(* Logix 5000 project; controller Joltek_RA_5069PLC002 vendor 1 type 14 code 226 rev 34.15; software revision 34.04 *)

TASK MainTask (continuous, watchdog 500 ms) : MainProgram
TASK SafetyTask (periodic, rate 20 ms, priority 10, watchdog 20 ms, safety) : SafetyProgram

MODULES
   Local : vendor 1 type 14 code 226 (5069 0, rev 34.15)
      Joltek_SW001 : vendor 1 type 12 code 231 (Ethernet 192.168.1.70, rev 13.8, Output RPI 1000 ms)
END_MODULES

TYPE UDT_ErrorDataLog :
STRUCT
   Time : UDT_Timestamp;
   DINTlog : DINT[10];
   REALlog : REAL[10];
END_STRUCT
END_TYPE

TYPE UDT_Timestamp :
STRUCT
   Year : DINT;
   Month : DINT;
   Day : DINT;
   Hour : DINT;
   Minute : DINT;
   Second : DINT;
END_STRUCT
END_TYPE

VAR_GLOBAL   (* controller tags *)
   Line34Pump3Motor342DischargeOfTank23_Sig : DINT;
   Line45Pump3MTR345InfeedRawIngredientFlou : DINT;
   Line6Pump1DischargeOfTank3 : DINT;
   Sys_DINT : DINT[100] := ([0] := 8, [1] := 1873, [2] := 997, [3] := 4, [5] := 10000, [6] := 10000, [39] := 50, [40] := 52, [41] := 6400, [42] := 3);
        [0]   // Line 1 Motor 324 of the Conveyor 23 Discharge Pump 4-20mA Signal
        [1]   // Line 2 Motor 32334 of the Conveyor 2233 Discharge Pump 0-20mA Signal SCALED
        [3].0   // Filler - Start
        [3].1   // Filler - Stop
        [3].3   // Filler - Faulted
        [3].2   // Filler - Running
        [4]   // Filler - Infeed Empty Bottle Count
        [40].4   // Capper - Start Capping Process
   Sys_FIFO_C : CONTROL[10] := ([0].LEN := 32, [0].POS := 2);
   Sys_Timer : TIMER[100] := ([0].PRE := 50, [0].ACC := 40, [0].EN := 1, [0].TT := 1, [1].PRE := 150, [1].ACC := 90, [1].EN := 1, [1].TT := 1, [2].PRE := 2000, [2].ACC := 184, [2].EN := 1, [2].TT := 1, [3].PRE := 200, [3].ACC := 136, [3].EN := 1, [3].TT := 1, [4].PRE := 200, [4].ACC := 162, [4].EN := 1, [4].TT := 1, [10].PRE := 200, [10].ACC := 147, [10].EN := 1, [10].TT := 1);
   System_Date_Time : DINT[7] := ([0] := 2025, [1] := 12, [2] := 8, [3] := 21, [4] := 13, [5] := 20, [6] := 843625);
   Test_Bool : BOOL[64];
END_VAR

PROGRAM MainProgram   (* main routine MainRoutine *)
VAR
   CurrentPos1 : DINT := 12;
END_VAR

ROUTINE _01_System   (* ladder *)
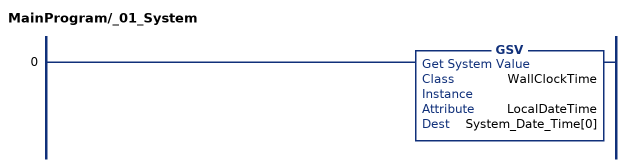
   0: GSV(WallClockTime,,LocalDateTime,System_Date_Time[0]);
END_ROUTINE

ROUTINE _02_Filler   (* ladder *)
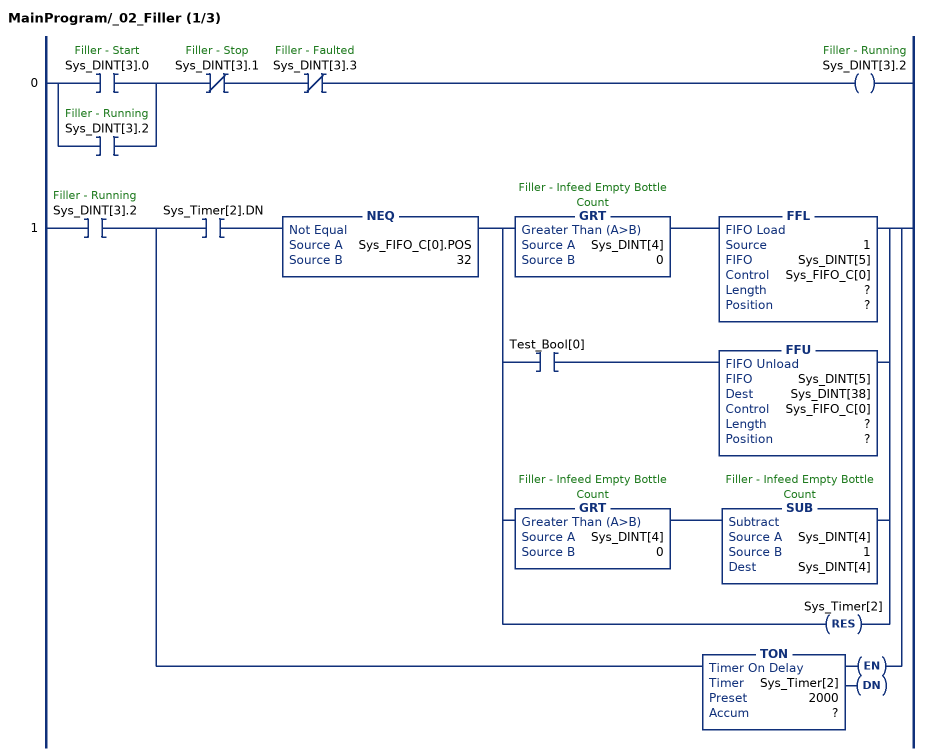
   0: [XIC(Sys_DINT[3].0) ,XIC(Sys_DINT[3].2) ]XIO(Sys_DINT[3].1)XIO(Sys_DINT[3].3)OTE(Sys_DINT[3].2);
   1: XIC(Sys_DINT[3].2)[XIC(Sys_Timer[2].DN) NEQ(Sys_FIFO_C[0].POS,32) [GRT(Sys_DINT[4],0) FFL(1,Sys_DINT[5],Sys_FIFO_C[0],?,?) ,XIC(Test_Bool[0]) FFU(Sys_DINT[5],Sys_DINT[38],Sys_FIFO_C[0],?,?) ,GRT(Sys_DINT[4],0) SUB(Sys_DINT[4],1,Sys_DINT[4]) ,RES(Sys_Timer[2]) ] ,TON(Sys_Timer[2],?,?) ];
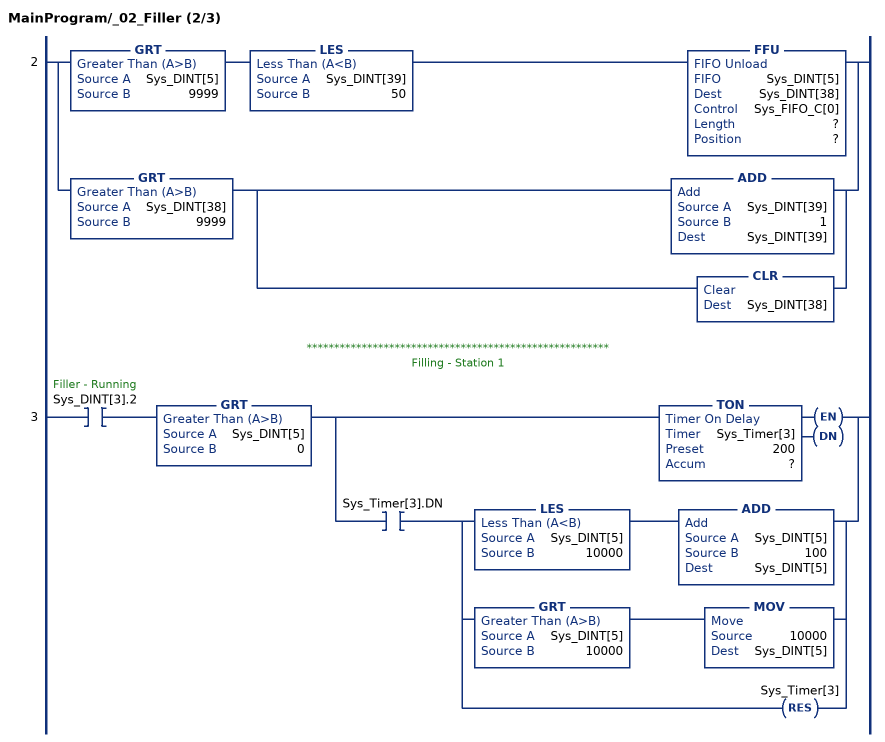
   2: [GRT(Sys_DINT[5],9999) LES(Sys_DINT[39],50) FFU(Sys_DINT[5],Sys_DINT[38],Sys_FIFO_C[0],?,?) ,GRT(Sys_DINT[38],9999) [ADD(Sys_DINT[39],1,Sys_DINT[39]) ,CLR(Sys_DINT[38]) ] ];
   // *******************************************************
   // Filling - Station 1
   3: XIC(Sys_DINT[3].2)GRT(Sys_DINT[5],0)[TON(Sys_Timer[3],?,?) ,XIC(Sys_Timer[3].DN) [LES(Sys_DINT[5],10000) ADD(Sys_DINT[5],100,Sys_DINT[5]) ,GRT(Sys_DINT[5],10000) MOV(10000,Sys_DINT[5]) ,RES(Sys_Timer[3]) ] ];
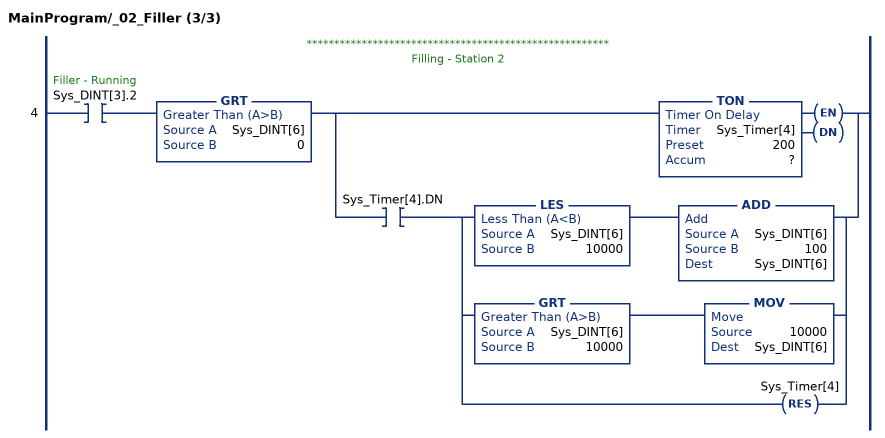
   // *******************************************************
   // Filling - Station 2
   4: XIC(Sys_DINT[3].2)GRT(Sys_DINT[6],0)[TON(Sys_Timer[4],?,?) ,XIC(Sys_Timer[4].DN) [LES(Sys_DINT[6],10000) ADD(Sys_DINT[6],100,Sys_DINT[6]) ,GRT(Sys_DINT[6],10000) MOV(10000,Sys_DINT[6]) ,RES(Sys_Timer[4]) ] ];
END_ROUTINE

ROUTINE _03_Capper   (* ladder *)
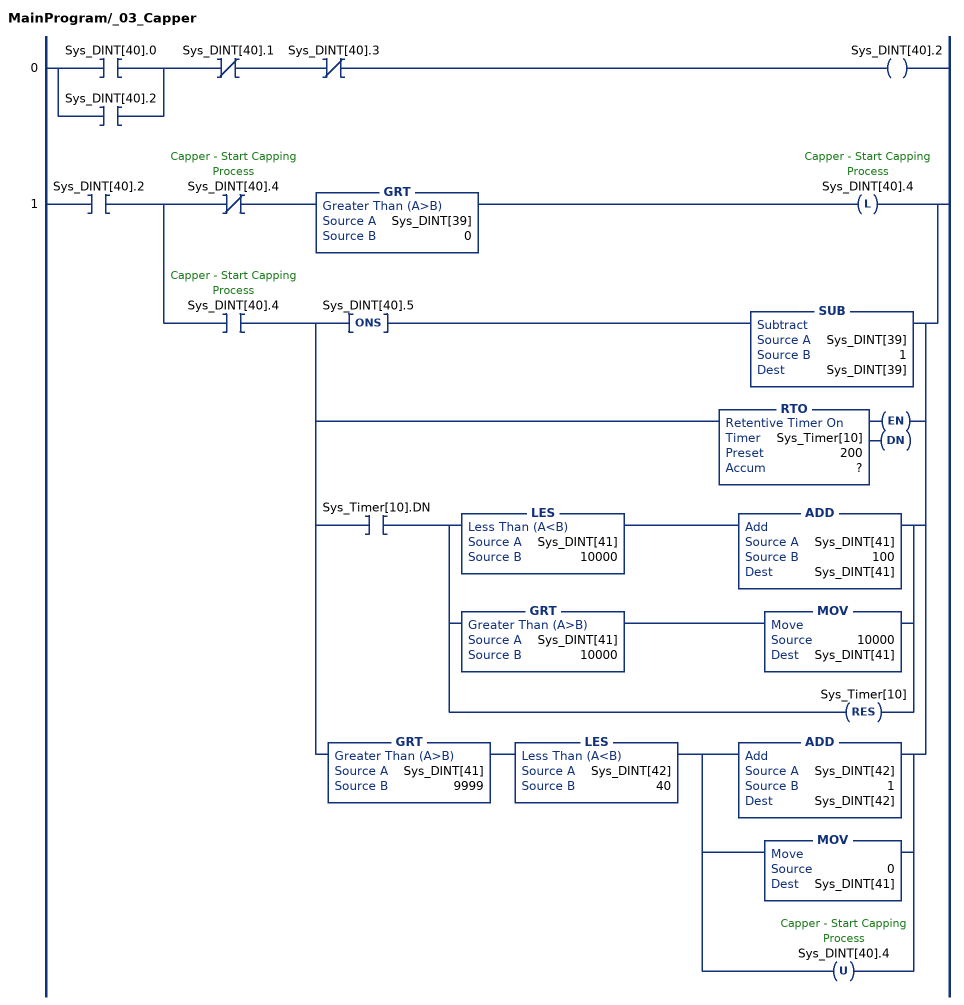
   0: [XIC(Sys_DINT[40].0) ,XIC(Sys_DINT[40].2) ]XIO(Sys_DINT[40].1)XIO(Sys_DINT[40].3)OTE(Sys_DINT[40].2);
   1: XIC(Sys_DINT[40].2)[XIO(Sys_DINT[40].4) GRT(Sys_DINT[39],0) OTL(Sys_DINT[40].4) ,XIC(Sys_DINT[40].4) [ONS(Sys_DINT[40].5) SUB(Sys_DINT[39],1,Sys_DINT[39]) ,RTO(Sys_Timer[10],?,?) ,XIC(Sys_Timer[10].DN) [LES(Sys_DINT[41],10000) ADD(Sys_DINT[41],100,Sys_DINT[41]) ,GRT(Sys_DINT[41],10000) MOV(10000,Sys_DINT[41]) ,RES(Sys_Timer[10]) ] ,GRT(Sys_DINT[41],9999) LES(Sys_DINT[42],40) [ADD(Sys_DINT[42],1,Sys_DINT[42]) ,MOV(0,Sys_DINT[41]) ,OTU(Sys_DINT[40].4) ] ] ];
END_ROUTINE

ROUTINE _04_Labeler   (* ladder *)
END_ROUTINE

ROUTINE _05_CasePacker   (* ladder *)
END_ROUTINE

ROUTINE _06_Palletizer   (* ladder *)
END_ROUTINE

ROUTINE _98_RandomizerLogic   (* ladder *)
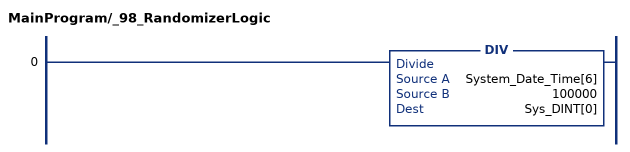
   0: DIV(System_Date_Time[6],100000,Sys_DINT[0]);
END_ROUTINE

ROUTINE _99_TestLogic   (* ladder *)
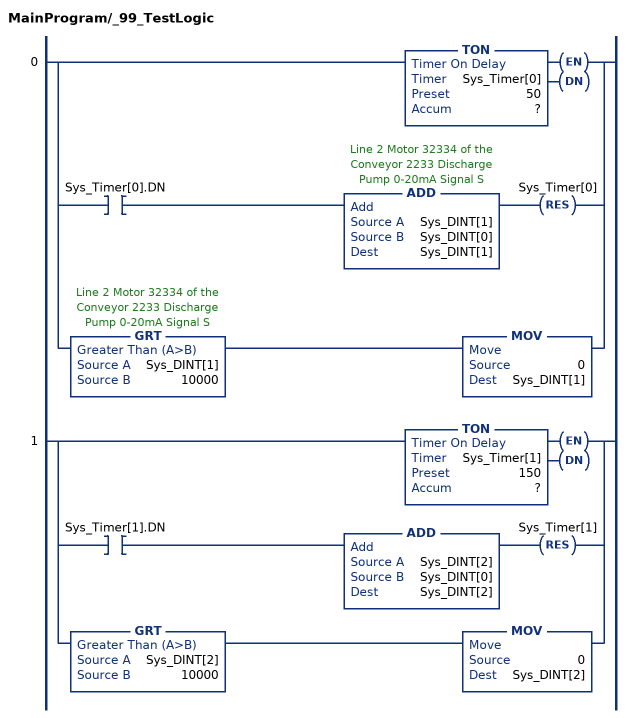
   0: [TON(Sys_Timer[0],?,?) ,XIC(Sys_Timer[0].DN) ADD(Sys_DINT[1],Sys_DINT[0],Sys_DINT[1]) RES(Sys_Timer[0]) ,GRT(Sys_DINT[1],10000) MOV(0,Sys_DINT[1]) ];
   1: [TON(Sys_Timer[1],?,?) ,XIC(Sys_Timer[1].DN) ADD(Sys_DINT[2],Sys_DINT[0],Sys_DINT[2]) RES(Sys_Timer[1]) ,GRT(Sys_DINT[2],10000) MOV(0,Sys_DINT[2]) ];
END_ROUTINE

ROUTINE MainRoutine   (* ladder *)
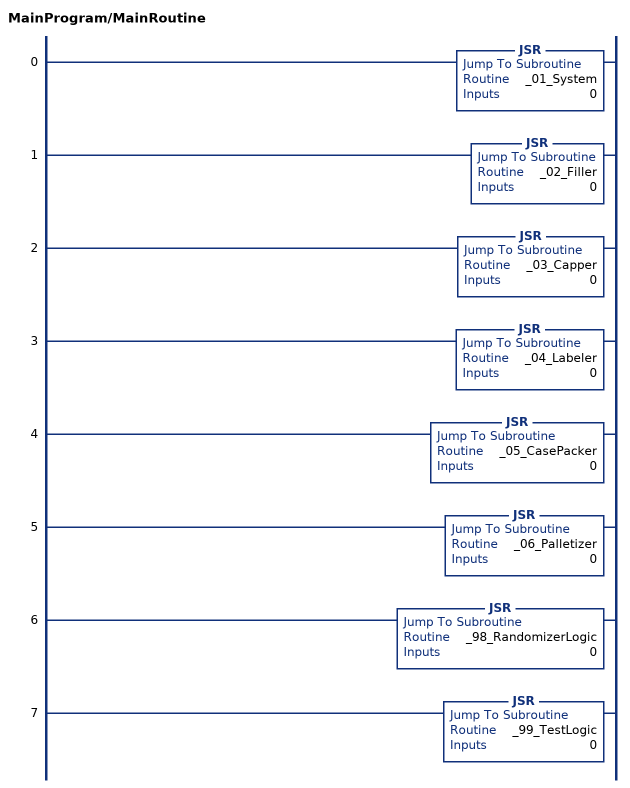
   0: JSR(_01_System,0);
   1: JSR(_02_Filler,0);
   2: JSR(_03_Capper,0);
   3: JSR(_04_Labeler,0);
   4: JSR(_05_CasePacker,0);
   5: JSR(_06_Palletizer,0);
   6: JSR(_98_RandomizerLogic,0);
   7: JSR(_99_TestLogic,0);
END_ROUTINE
END_PROGRAM

PROGRAM SafetyProgram   (* main routine MainRoutine, safety *)

ROUTINE MainRoutine   (* ladder *)
END_ROUTINE
END_PROGRAM
